
     // Eleminate "third" coordinate
     CASE #pathPlane OF
       "CP_XY":
         #tempVectorA.z := 0.0;
         #tempVectorB.z := 0.0;

       "CP_XZ":
         #tempVectorA.y := 0.0;
         #tempVectorB.y := 0.0;

       "CP_YZ":
         #tempVectorA.x := 0.0;
         #tempVectorB.x := 0.0;
     END_CASE;

     #distancePathPlane := "LKinCtrl_VecAbs"("LKinCtrl_VecSub"(vIn1:=#tempVectorB, vIn2:=#tempVectorA));



   END_REGION CALCULATION

   #LKinCtrl_CalcVecDistancePathPlane := 0; // o.k.
END_FUNCTION

FUNCTION "LKinCtrl_CalcToolLengthCompensation" : Word   // FC35070, SCL
TITLE = LKinCtrl_CalcToolLengthCompensation
{ S7_Optimized_Access := 'TRUE' }
AUTHOR : tech.team.motioncontrol@siemens.com
FAMILY : LKinCtrl
VERSION : 1.0
// Calculate tool length compensation according to path plane and absolute / relative
   VAR_INPUT
      toolLength : LReal;   // Tool length
      pathPlane : Int;   // Path plane: XZ= 0, YZ=1, XY= 2
   END_VAR
   VAR_IN_OUT
      point : "LKinCtrl_typeCOff3DPoint";   // PositioningAxis to get data from
   END_VAR
   // Ret_Val : Return value
   VAR CONSTANT
      ERR_COFF_INVALID_PATH_PLANE : Word := 16#8303;   // Error - invalid path plane
   END_VAR
BEGIN
   //=============================================================================
   // SIEMENS AG
   // (c)Copyright 2019 All Rights Reserved
   //-----------------------------------------------------------------------------
   // Library: - 
   // Tested with: S7-1516T-3 PN
   // Engineering: TIA Portal V15
   // Restrictions: -
   // Requirements: S7-1500/S7-1500T FW 2.5
   // Functionality: Calculate tool length compensation according to path plane and absolute / relative
   // Result ist the compensated coordinate
   // and end point
   //-----------------------------------------------------------------------------
   // Change log table:
   // Version  Date       Expert in charge Changes applied
   // 01.00.00 2019-02-11 AW               created
   //=============================================================================

   REGION PLAUSIBILITY_CHECK
   // Check path plane
   IF ((#pathPlane >= "CP_XZ") AND (#pathPlane <= "CP_XY"))
   THEN
     ;
   ELSE
     #LKinCtrl_CalcToolLengthCompensation := #ERR_COFF_INVALID_PATH_PLANE; // Invalid path plane
     RETURN;
   END_IF;
   END_REGION PLAUSIBILITY_CHECK

   REGION CALCULATION

     CASE #pathPlane OF
       "CP_XY":
         #point.z += #toolLength;
       "CP_XZ":
         #point.y += #toolLength;
       "CP_YZ":
         #point.x += #toolLength;
     END_CASE;


   END_REGION CALCULATION

   #LKinCtrl_CalcToolLengthCompensation := 0; // o.k.
END_FUNCTION

FUNCTION "LKinCtrl_VecAdd" : "LKinCtrl_typeCOff3DPoint"   // FC35080, SCL
TITLE = LKinCtrl_VecAdd
{ S7_Optimized_Access := 'TRUE' }
AUTHOR : tech.team.motioncontrol@siemens.com
FAMILY : LKinCtrl
VERSION : 1.0
// Add two coordinates (X, Y, Z) of "LKinCtrl_typeCOff3DPoint"
   VAR_INPUT
      vIn1 : "LKinCtrl_typeCOff3DPoint";   // Input vector 1
      vIn2 : "LKinCtrl_typeCOff3DPoint";   // Input vector 2
   END_VAR
   // Ret_Val : Return value - calculated vector
BEGIN
   //=============================================================================
   // SIEMENS AG
   // (c)Copyright 2018 All Rights Reserved
   //-----------------------------------------------------------------------------
   // Library: - 
   // Tested with: S7-1516T-3 PN
   // Engineering: TIA Portal V15
   // Restrictions: -
   // Requirements: S7-1500/S7-1500T FW 2.5
   // Functionality: Add two coordinates (X, Y, Z) of "LKinCtrl_typeCOff3DPoint"
   //-----------------------------------------------------------------------------
   // Change log table:
   // Version  Date       Expert in charge Changes applied
   // 01.00.00 2018-10-26 AW               created
   //=============================================================================
   #LKinCtrl_VecAdd.x := #vIn1.x + #vIn2.x;
   #LKinCtrl_VecAdd.y := #vIn1.y + #vIn2.y;
   #LKinCtrl_VecAdd.z := #vIn1.z + #vIn2.z;
END_FUNCTION

FUNCTION "LKinCtrl_VecSub" : "LKinCtrl_typeCOff3DPoint"   // FC35081, SCL
TITLE = LKinCtrl_VecSub
{ S7_Optimized_Access := 'TRUE' }
AUTHOR : tech.team.motioncontrol@siemens.com
FAMILY : LKinCtrl
VERSION : 1.0
// Substract two coordinates (X, Y, Z) of "LKinCtrl_typeCOff3DPoint"
   VAR_INPUT
      vIn1 : "LKinCtrl_typeCOff3DPoint";   // Input vector 1
      vIn2 : "LKinCtrl_typeCOff3DPoint";   // Input vector 2
   END_VAR
   // Ret_Val : Return value - difference vector
BEGIN
   //=============================================================================
   // SIEMENS AG
   // (c)Copyright 2018 All Rights Reserved
   //-----------------------------------------------------------------------------
   // Library: - 
   // Tested with: S7-1516T-3 PN
   // Engineering: TIA Portal V15
   // Restrictions: -
   // Requirements: S7-1500/S7-1500T FW 2.5
   // Functionality: Substract two coordinates (X, Y, Z) of "LKinCtrl_typeCOff3DPoint"
   //-----------------------------------------------------------------------------
   // Change log table:
   // Version  Date       Expert in charge Changes applied
   // 01.00.00 2018-10-26 AW               created
   //=============================================================================
   #LKinCtrl_VecSub.x := #vIn1.x - #vIn2.x;
   #LKinCtrl_VecSub.y := #vIn1.y - #vIn2.y;
   #LKinCtrl_VecSub.z := #vIn1.z - #vIn2.z;
END_FUNCTION

FUNCTION "LKinCtrl_VecUnit" : "LKinCtrl_typeCOff3DPoint"   // FC35082, SCL
TITLE = LKinCtrl_VecUnit
{ S7_Optimized_Access := 'TRUE' }
AUTHOR : tech.team.motioncontrol@siemens.com
FAMILY : LKinCtrl
VERSION : 1.0
// Create unit vector of coordinates (X, Y, Z) of "LKinCtrl_typeCOff3DPoint"
   VAR_INPUT
      vIn : "LKinCtrl_typeCOff3DPoint";   // Input vector
   END_VAR
   // Ret_Val : Return value - unit vector
BEGIN
   //=============================================================================
   // SIEMENS AG
   // (c)Copyright 2018 All Rights Reserved
   //-----------------------------------------------------------------------------
   // Library: - 
   // Tested with: S7-1516T-3 PN
   // Engineering: TIA Portal V15
   // Restrictions: -
   // Requirements: S7-1500/S7-1500T FW 2.5
   // Functionality: Create unit vector of coordinates (X, Y, Z) of "LKinCtrl_typeCOff3DPoint"
   //-----------------------------------------------------------------------------
   // Change log table:
   // Version  Date       Expert in charge Changes applied
   // 01.00.00 2018-08-27 SF               created
   //=============================================================================

   //Out = In/abs(In)
   #LKinCtrl_VecUnit := "LKinCtrl_VecDivScal"(vIn := #vIn,
                                              sIn := "LKinCtrl_VecAbs"(#vIn));
END_FUNCTION

FUNCTION "LKinCtrl_VecAbs" : LReal   // FC35083, SCL
TITLE = LKinCtrl_VecAbs
{ S7_Optimized_Access := 'TRUE' }
AUTHOR : tech.team.motioncontrol@siemens.com
FAMILY : LKinCtrl
VERSION : 1.0
// Calculate length of vector of coordinates (X, Y, Z) of "LKinCtrl_typeCOff3DPoint"
   VAR_INPUT
      vIn : "LKinCtrl_typeCOff3DPoint";   // Input vector
   END_VAR
   // Ret_Val : Return value - scalar
BEGIN
   //=============================================================================
   // SIEMENS AG
   // (c)Copyright 2018 All Rights Reserved
   //-----------------------------------------------------------------------------
   // Library: - 
   // Tested with: S7-1516T-3 PN
   // Engineering: TIA Portal V15
   // Restrictions: -
   // Requirements: S7-1500/S7-1500T FW 2.5
   // Functionality: Calculate length of vector of coordinates (X, Y, Z) of "LKinCtrl_typeCOff3DPoint"
   //-----------------------------------------------------------------------------
   // Change log table:
   // Version  Date       Expert in charge Changes applied
   // 01.00.00 2018-10-26 AW               created
   //=============================================================================

   #LKinCtrl_VecAbs := SQRT(#vIn.x*#vIn.x + #vIn.y*#vIn.y + #vIn.z*#vIn.z);
END_FUNCTION

FUNCTION "LKinCtrl_VecScale" : "LKinCtrl_typeCOff3DPoint"   // FC35084, SCL
TITLE = LKinCtrl_VecScale
{ S7_Optimized_Access := 'TRUE' }
AUTHOR : tech.team.motioncontrol@siemens.com
FAMILY : LKinCtrl
VERSION : 1.0
// Scale vector (X, Y, Z) of "LKinCtrl_typeCOff3DPoint"
   VAR_INPUT
      vIn : "LKinCtrl_typeCOff3DPoint";   // Input vector
      factor : LReal;   // Scaling factor
   END_VAR
   // Ret_Val : Return value - scaled vector
BEGIN
   //=============================================================================
   // SIEMENS AG
   // (c)Copyright 2018 All Rights Reserved
   //-----------------------------------------------------------------------------
   // Library: - 
   // Tested with: S7-1516T-3 PN
   // Engineering: TIA Portal V15
   // Restrictions: -
   // Requirements: S7-1500/S7-1500T FW 2.5
   // Functionality: Scale vector (X, Y, Z) of "LKinCtrl_typeCOff3DPoint"
   //-----------------------------------------------------------------------------
   // Change log table:
   // Version  Date       Expert in charge Changes applied
   // 01.00.00 2018-10-26 AW               created
   //=============================================================================

   #LKinCtrl_VecScale.x := #vIn.x * #factor;
   #LKinCtrl_VecScale.y := #vIn.y * #factor;
   #LKinCtrl_VecScale.z := #vIn.z * #factor;
END_FUNCTION

FUNCTION "LKinCtrl_VecDivScal" : "LKinCtrl_typeCOff3DPoint"   // FC35085, SCL
TITLE = LKinCtrl_VecDivScal
{ S7_Optimized_Access := 'TRUE' }
AUTHOR : tech.team.motioncontrol@siemens.com
FAMILY : LKinCtrl
VERSION : 1.0
// Divide coordinate with scalar of coordinates (X, Y, Z) of "LKinCtrl_typeCOff3DPoint"
   VAR_INPUT
      vIn : "LKinCtrl_typeCOff3DPoint";   // Input vector
      sIn : LReal;   // Input scalar
   END_VAR
   // Ret_Val : Return value - calculated vector
BEGIN
   //=============================================================================
   // SIEMENS AG
   // (c)Copyright 2018 All Rights Reserved
   //-----------------------------------------------------------------------------
   // Library: - 
   // Tested with: S7-1516T-3 PN
   // Engineering: TIA Portal V15
   // Restrictions: -
   // Requirements: S7-1500/S7-1500T FW 2.5
   // Functionality: Divide coordinate with scalar of coordinates (X, Y, Z) of "LKinCtrl_typeCOff3DPoint"
   //-----------------------------------------------------------------------------
   // Change log table:
   // Version  Date       Expert in charge Changes applied
   // 01.00.00 2018-10-26 AW               created
   //=============================================================================

   IF (#sIn <> 0.0) THEN
     #LKinCtrl_VecDivScal.x := #vIn.x / #sIn;
     #LKinCtrl_VecDivScal.y := #vIn.y / #sIn;
     #LKinCtrl_VecDivScal.z := #vIn.z / #sIn;
   ELSE
     #LKinCtrl_VecDivScal.x := 0.0;
     #LKinCtrl_VecDivScal.y := 0.0;
     #LKinCtrl_VecDivScal.z := 0.0;
   END_IF;
END_FUNCTION

FUNCTION "LKinCtrl_VecScalProd" : LReal   // FC35086, SCL
TITLE = LKinCtrl_VecScalProd
{ S7_Optimized_Access := 'TRUE' }
AUTHOR : tech.team.motioncontrol@siemens.com
FAMILY : LKinCtrl
VERSION : 1.0
// Calculate scalar product of coordinates (X, Y, Z) of "LKinCtrl_typeCOff3DPoint"
   VAR_INPUT
      vIn1 : "LKinCtrl_typeCOff3DPoint";   // Input vector 1
      vIn2 : "LKinCtrl_typeCOff3DPoint";   // Input vector 2
   END_VAR
   // Ret_Val : Scalar product
BEGIN
   //=============================================================================
   // SIEMENS AG
   // (c)Copyright 2019 All Rights Reserved
   //-----------------------------------------------------------------------------
   // Library: - 
   // Tested with: S7-1516T-3 PN
   // Engineering: TIA Portal V15
   // Restrictions: -
   // Requirements: S7-1500/S7-1500T FW 2.5
   // Functionality: Calculate scalar product of coordinates (X, Y, Z) of "LKinCtrl_typeCOff3DPoint"
   //-----------------------------------------------------------------------------
   // Change log table:
   // Version  Date       Expert in charge Changes applied
   // 01.00.00 2019-01-25 AW               created
   //=============================================================================

   #LKinCtrl_VecScalProd := #vIn1.x * #vIn2.x  //   X1*X2
                          + #vIn1.y * #vIn2.y  // + Y1*Y2
                          + #vIn1.z * #vIn2.z; // + Z1*Z2
END_FUNCTION

FUNCTION "LKinCtrl_VecCrossProd" : "LKinCtrl_typeCOff3DPoint"   // FC35087, SCL
TITLE = LKinCtrl_VecCrossProd
{ S7_Optimized_Access := 'TRUE' }
AUTHOR : tech.team.motioncontrol@siemens.com
FAMILY : LKinCtrl
VERSION : 1.0
// Cross product of two coordinates (X, Y, Z) of "LKinCtrl_typeCOff3DPoint"
   VAR_INPUT
      vIn1 : "LKinCtrl_typeCOff3DPoint";   // Input vector 1
      vIn2 : "LKinCtrl_typeCOff3DPoint";   // Input vector 2
   END_VAR
   // Ret_Val : Return value - calculated vector
BEGIN
   //=============================================================================
   // SIEMENS AG
   // (c)Copyright 2018 All Rights Reserved
   //-----------------------------------------------------------------------------
   // Library: - 
   // Tested with: S7-1516T-3 PN
   // Engineering: TIA Portal V15
   // Restrictions: -
   // Requirements: S7-1500/S7-1500T FW 2.5
   // Functionality: Cross product of two coordinates (X, Y, Z) of "LKinCtrl_typeCOff3DPoint"
   //-----------------------------------------------------------------------------
   // Change log table:
   // Version  Date       Expert in charge Changes applied
   // 01.00.00 2019-01-24 AW               created
   //=============================================================================

   #LKinCtrl_VecCrossProd.x := #vIn1.y * #vIn2.z - #vIn1.z * #vIn2.y;
   #LKinCtrl_VecCrossProd.y := #vIn1.z * #vIn2.x - #vIn1.x * #vIn2.z;
   #LKinCtrl_VecCrossProd.z := #vIn1.x * #vIn2.y - #vIn1.y * #vIn2.x;
END_FUNCTION

// folder: LKinCtrl_Blocks/LKinCtrl_SubBlocks/LKinCtrl_SubCalcBlocks

FUNCTION_BLOCK "LKinCtrl_SetFlagCtrl"   // FB35024, SCL
TITLE = LKinCtrl_SetFlagCtrl / Enable Template
{ S7_Optimized_Access := 'TRUE' }
AUTHOR : tech.team.motioncontrol@siemens.com
FAMILY : LKinCtrl
VERSION : 2.0
// Handle setFlags in FB MovePath / Template for an FB with Enable / Valid handling based on PLCopen standard "Function Blocks for Motion Control" V2.0
   VAR_INPUT
      enable : Bool;   // TRUE: Enable functionality of FB
      activeCmdNo : DInt;   // Number of actual PathData set number (interconnect LKinCtrl_MC_ExecuteKinMotionCmd)
      activePathDataIdentifier : USInt;   // Identifier number of actual PathData (interconnect LKinCtrl_MC_ExecuteKinMotionCmd)
      activePathDataName : String["LKINCTRL_LENGTH_OF_PATHDATA_NAME"];   // Name of actual PathData (interconnect LKinCtrl_MC_ExecuteKinMotionCmd)
      remainingDistanceActCmd : LReal;   // RemainingDistance of active motionCommand (interconnect LKinCtrl_MC_ExecuteKinMotionCmd)
      kinematicsStatusWord : DWord;   // Interconnect axesGroup.StatusWord / Interconnect 'axesGroup.StatusWord.X9'
      movePathStatus : Word;   // Interconnect value for MovePath output 'status'
      flagsBuffer : Struct   // Buffer to store flag information for past and actual commands
         writeBufferElement : Int := 1;   // pointer on entry to be written
         bufferElement : Array[1.."LKINCTRL_NO_OF_SETFLAGS_BUFFER_ELEMENTS"] of Struct   // flag information for one specific command (see cmdId)
            pathDataName : String["LKINCTRL_LENGTH_OF_PATHDATA_NAME"];   // PathData name of specific command
            pathDataIdentifier : DInt;   // PathData identifier counter of specific command
            cmdId : DInt;   // cmdId of command in PathData
            isIntermediateCmd : Bool;   // TRUE: command is intermediate command
            setFlags : Array[1.."LKINCTRL_NO_OF_CMD_SETFLAGS"] of "LKinCtrl_typeSetFlagElement_Bool";   // setFlags structure equal to PathData command entry
            valueFlags : Array[1.."LKINCTRL_NO_OF_CMD_VALUEFLAGS"] of "LKinCtrl_typeSetFlagElement_LReal";   // setFlags structure equal to PathData command entry
         END_STRUCT;
      END_STRUCT;
   END_VAR
   VAR_OUTPUT
      valid : Bool;   // TRUE: Valid set of output values available at the FB
      busy : Bool;   // TRUE: FB is not finished and new output values can be expected
      error : Bool;   // TRUE: An error occurred during the execution of the FB
      status : Word := 16#7000;   // 16#0000 - 16#7FFF: Status of the FB, 16#8000 - 16#FFFF: Error identification
      waitMain : Bool;   // Static bit to wait for execution due to wait flags & valueFlags
   END_VAR
   VAR_IN_OUT
      flags : Array[0.."LKINCTRL_NO_OF_LAST_SETFLAG"] of Bool;   // Interconnect MovePath outputs for flag signals
      waitFlags : Struct   // Static struct to store wait flag information
         waitCtr : Int;   // counter for number of wait flags in one command
         waitFlag : Array[1.."LKINCTRL_NO_OF_CMD_SETFLAGS"] of Int;   // flag number as identifier for flag active as wait flag
      END_STRUCT;
   END_VAR
   VAR
      statEnableOld : Bool;   // Old value of 'enable' input for edge detection
      statValid : Bool;   // Static value for output 'valid'
      statBusy : Bool;   // Static value for output 'busy'
      statError : Bool;   // Static value for output 'error'
      statErrorUserCleared : Bool;   // Error occurred that can only be solved by user; rising edge at enable input necessary
      statErrorAutoCleared : Bool;   // Error occurred that can be acknowledged by FB
      statStatus : Word := 16#7000;   // Static value for output 'status'
      statFBState : DInt := 0;   // State in the state machine of the FB
      statDisablingCompleted : Bool;   // TRUE: Disabling has been completed
      statWaitMain : Bool;   // Static value for output 'waitMain'
      statSkippedCmdCounter : Int;   // Static counter for skipped activeCmdNo
      statActivePathDataIdentifierOld : USInt;   // Static to store old activePathDataIdentifier from LKinCtrl_ExecuteKinMotionCmd
      statActiveCmdNoOld : DInt;   // Static variable storing old 'activeCmdNo'
      statActivePathDataNameOld : String["LKINCTRL_LENGTH_OF_PATHDATA_NAME"];   // Static to store last active PathData name
      statFlagSetAfterCmd : Array[1.."LKINCTRL_NO_OF_CMD_SETFLAGS"] of Int;   // Static array storing flags to be set after command
      statWaitFlagSetAfterCmd : Array[1.."LKINCTRL_NO_OF_CMD_SETFLAGS"] of Int;   // Static array storing wait flags to be set after command / Static array storing flags to be set after command
      statFlagResetAfterOneCmd : Array[1.."LKINCTRL_NO_OF_CMD_SETFLAGS"] of Int;   // Static array storing flags to be reset after one command
      statFlagResetFM3 : Array[1.."LKINCTRL_NO_OF_CMD_SETFLAGS"] of Int;   // Static array storing flags to be reset after one cycle
      statFlagSetFM10 : Array[1.."LKINCTRL_NO_OF_CMD_SETFLAGS"] of Int;   // Static array storing flags to be set at remaining distance
      statRemDistanceFM10 : Array[1.."LKINCTRL_NO_OF_CMD_SETFLAGS"] of LReal;   // Static array storing remaining distance for flags
      statFlagSetFM13 : Array[1.."LKINCTRL_NO_OF_CMD_SETFLAGS"] of Int;   // Static array storing flags to be set after command for one cycle
      statFlagResetFM13 : Array[1.."LKINCTRL_NO_OF_CMD_SETFLAGS"] of Int;   // Static array storing flags to be set after command and reset after one cycle
      statWaitFlagActiveCmdId : Array[1.."LKINCTRL_NO_OF_CMD_SETFLAGS"] of DInt;   // Static array storing active command number for watiFlag
      statWaitFlagActivePathData : Array[1.."LKINCTRL_NO_OF_CMD_SETFLAGS"] of DInt;   // Static array storing active PathData number for watiFlag
      statFlagResetSkipped : Array[1..#MAX_NUMBER_OF_SKIPPED_CMDS, 1.."LKINCTRL_NO_OF_CMD_SETFLAGS"] of Int;   // Static array storing flags to be reset after one cycle
      statWaitFlagOld : Array[1.."LKINCTRL_NO_OF_CMD_SETFLAGS"] of Bool;   // Static array storing last flag values for reset detection
   END_VAR
   VAR_TEMP
      tempEnable : Bool;   // Temporary value for input 'enable'
      tempFlagCmdCounter : Int;   // Temporary flag cmd counter for setFlag UDT
      tempFlagsBufferElementCtr : Int;   // Temporary flag buffer counter
      tempFlagCounter : Int;   // Temporary flag counter for flag array
      tempFlagWasSet : Bool;   // Temporary bool to signalize flag was set after end of PRG
      tempSkippedCounterInc : Bool;   // Temporary bool to signalize skipped counter was increased
   END_VAR
   VAR CONSTANT
      FB_STATE_NO_PROCESSING : DInt := 0;   // FB state: No processing
      FB_STATE_CHECK_ACTIVE_CMD : DInt := 50;   // FB state: Check change of active command
      FB_STATE_SET_RESET_AFTER_COMMAND : DInt := 51;   // FB state: Handle flag actions after commands
      FB_STATE_EVALUATE_FLAGBUFFER : DInt := 52;   // FB state: Handle flagBuffer and flag actions before command
      FB_STATE_RESET_AFTER_ONE_CYCLE : DInt := 53;   // FB state: Handle flag reset after one cycle
      FB_STATE_CHECK_REMAINING_DISTANCE : DInt := 54;   // FB state: Check flag with remaining distance
      FB_STATE_WAIT_FLAG_HANDLING : DInt := 55;   // FB state: Check wait flags
      FB_STATE_DISABLING : DInt := 90;   // FB state: Disabling
      STATUS_NO_CALL : Word := 16#7000;   // No job being currently processed
      STATUS_FIRST_CALL : Word := 16#7001;   // First call after incoming new job (rising edge 'execute')
      STATUS_SUBSEQUENT_CALL : Word := 16#7002;   // Subsequent call during active processing without further details
      ERR_UNDEFINED_STATE : Word := 16#8600;   // Error due to an undefined state in state machine
      ERR_OVERFLOW_SKIPPED_CMDS : Word := 16#8601;   // Error due to overflow of skipped commands counter
      STATUS_EXECUTION_WAITING : Word := 16#7307;   // Status path execution waiting due to wait flag, wait time or single step mode
      MAX_NUMBER_OF_SKIPPED_CMDS : Int := 3;   // Maximum number of activeCmdNo to be skipped
      SPTP_REMAINING_DIST : Bool := FALSE;   // TRUE: Caclulate own RemainingDistance for SPTP / FALSE: Use ExecutionTimeStatus
   END_VAR
   // flagsBuffer.bufferElement[1].pathDataName := '';
   // flagsBuffer.bufferElement[1].cmdId := 0;
BEGIN
   //==========================================================================================
   // SIEMENS AG
   // (c)Copyright 2020 All Rights Reserved
   //------------------------------------------------------------------------------------------
   // Library: LKinCtrl
   // Tested with: S7-1517T-3 PN/DP
   // Engineering: TIA Portal V15
   // Restrictions: ---
   // Requirements: S7-1500T FW 2.5
   // Functionality: LKinCtrl_SetFlagCtrl
   // The FC evaluates the flag informaton given by the PathData structure and controls the flag
   // variables depending on the active command information given
   // 
   // Support: tech.team.motioncontrol@siemens.com
   // Note: Parameter comments are only available in language 'English (United States)'
   //------------------------------------------------------------------------------------------
   // Change log table:
   // Version    Date          Expert in charge    Changes applied
   // 01.00.00   19.08.2019    JR                  First release version v1.0
   // 01.00.01   18.09.2019    JR                  Updates for LREAL flags
   // 01.00.02   19.09.2019    JR                  Implementation wait value flags - flagMode 5
   // 01.00.03   19.09.2019    JR                  Implementation value flags - flagMode 11 - 15
   // 01.00.04   27.11.2019    JR                  Additional condition for deactivating flags
   // 01.01.00   28.11.2019    JR                  Separate block for setFlags from LKinCtrl_FlagCtrl
   // 01.01.01   27.01.2020    FR                  Changed FM 10 from > to >=
   // 01.01.02   30.01.2020    FR                  Changed flag array constant
   // 02.00.00   12.03.2020    FR                  Reworked complete FB to fit enable template with state machine
   // 02.00.01   17.03.2020    FR                  Check remDistance <= 0.0 instead of =
   // 02.00.02   03.08.2020    FR                  Change interface actualCmdIsCircularCmd to KinematicsStatusWord (DWord)
   // 02.00.03   19.10.2020    FR                  Handle multiple commands per cycle; Changed case to use constants instead of numbers
   // 02.00.04   15.12.2020    FR                  Added option for SPTP commands to have calculated remainingDistance
   // 02.00.05   01.06.2021    FR                  Use variable instead of F_Trig, Fix for FM5 / FM15, Fix for statActiveCmdNoOld not being reset correctly
   // 02.00.06   06.07.2021    FR                  Save old variables only when processed
   //===========================================================================================

   #tempEnable := #enable; // Work with temporary value / create process image

   REGION ENABLING/DISABLING
     IF (#tempEnable = TRUE) AND (#statStatus = #STATUS_NO_CALL) THEN // Enable FB
       // First call; initialize FB
       #statValid := TRUE;
       #statBusy := TRUE;
       #statError := FALSE;
       #statErrorUserCleared := FALSE;
       #statErrorAutoCleared := FALSE;
       #statStatus := #STATUS_FIRST_CALL;

       #statFBState := #FB_STATE_CHECK_ACTIVE_CMD; // State machine - start functionality
       //------------------------------------------------------------------------------------------
       // Initialize functionality: reset of variables, diagnostics, etc.
       #statDisablingCompleted := FALSE;

       // Initialize all setFlags (flag array) when enabling
       //------------------------------------------------------------------------------------------
       FOR #tempFlagCounter := 0 TO "LKINCTRL_NO_OF_LAST_SETFLAG" DO
         #flags[#tempFlagCounter] := FALSE;
       END_FOR;

       // Initialize flag handling variables
       //------------------------------------------------------------------------------------------
       // reset wait output
       #statWaitMain := FALSE;
       #statSkippedCmdCounter := 0;
       #statActiveCmdNoOld := 0;
       #statActivePathDataNameOld := '';
       #statActivePathDataIdentifierOld := 0;

       FOR #tempFlagCmdCounter := 1 TO "LKINCTRL_NO_OF_CMD_SETFLAGS" DO
         // reset auxiliary flag storage variables
         #statFlagResetAfterOneCmd[#tempFlagCmdCounter] := -1;
         #statFlagSetAfterCmd[#tempFlagCmdCounter] := -1;
         #statWaitFlagSetAfterCmd[#tempFlagCmdCounter] := -1;
         #statFlagResetFM3[#tempFlagCmdCounter] := -1;
         #statFlagResetFM13[#tempFlagCmdCounter] := -1;
         #statFlagSetFM13[#tempFlagCmdCounter] := -1;
         #statFlagSetFM10[#tempFlagCmdCounter] := -1;
         #statRemDistanceFM10[#tempFlagCmdCounter] := 0.0;
         #statWaitFlagActiveCmdId[#tempFlagCmdCounter] := 0;
         #statWaitFlagActivePathData[#tempFlagCmdCounter] := 0;

         // Initialize functionality: call subsidiary FBs with FALSE
         #statWaitFlagOld[#tempFlagCmdCounter] := FALSE;

         // Reset storage for skipped commands
         FOR #tempFlagCounter := 1 TO #MAX_NUMBER_OF_SKIPPED_CMDS DO
           #statFlagResetSkipped[#tempFlagCounter, #tempFlagCmdCounter] := -1;
         END_FOR;
       END_FOR;


       //------------------------------------------------------------------------------------------

     ELSIF (#tempEnable = FALSE) AND (#statEnableOld = TRUE) THEN // Disable FB 
       #statFBState := #FB_STATE_DISABLING;

     ELSIF (#statStatus = #STATUS_FIRST_CALL) THEN // Set status identifier of subsequent call
       #statStatus := #STATUS_SUBSEQUENT_CALL;
     END_IF;

     // Edge detection 'enable' input
     #statEnableOld := #tempEnable;
   END_REGION ENABLING/DISABLING

   IF (#statStatus = #STATUS_NO_CALL) THEN // Nothing to do -> End here to reduce "system load"
     RETURN;
   END_IF;

   REGION STATE_MACHINE
     // Use if sate machine for more states in one cycle

     // No processing active (Note: this state must always be present and left empty)
     IF #statFBState = #FB_STATE_NO_PROCESSING THEN
       ;
     END_IF;

     // Reset after one cycle 
     REGION STATE_RESET_AFTER_ONE_CYCLE
       IF #statFBState = #FB_STATE_RESET_AFTER_ONE_CYCLE THEN
         // for loop checking all available flags
         FOR #tempFlagCmdCounter := 1 TO "LKINCTRL_NO_OF_CMD_SETFLAGS" DO
           // reset flags active for one cycle only (flagMode: 3)
           IF #statFlagResetFM3[#tempFlagCmdCounter] <> -1 THEN
             // reset flags when active command is ended / next command starts
             #flags[#statFlagResetFM3[#tempFlagCmdCounter]] := FALSE;
             // reset stored flag to be reset (to not reset it after each single future command)
             #statFlagResetFM3[#tempFlagCmdCounter] := -1;
           END_IF;

           // reset flags active for one cycle only (flagMode: 13)
           IF #statFlagResetFM13[#tempFlagCmdCounter] <> -1 THEN
             // reset flags when active command is ended / next command starts
             #flags[#statFlagResetFM13[#tempFlagCmdCounter]] := FALSE;
             // reset stored flag to be reset (to not reset it after each single future command)
             #statFlagResetFM13[#tempFlagCmdCounter] := -1;
           END_IF;

           // Check if commands were skipped and reset flags
           FOR #tempFlagCounter := 1 TO #statSkippedCmdCounter DO // If no cmd was skipped the upper limit should be 0 --> No execution of the loop
             // If activeCmdNo was skipped reset flags active for one cycle only (flagMode: 2/3/13)
             IF #statFlagResetSkipped[#tempFlagCounter, #tempFlagCmdCounter] <> -1 THEN
               // reset flags when active command is ended / next command starts
               #flags[#statFlagResetSkipped[#tempFlagCounter, #tempFlagCmdCounter]] := FALSE;
               // reset stored flag to be reset (to not reset it after each single future command)
               #statFlagResetSkipped[#tempFlagCounter, #tempFlagCmdCounter] := -1;
             END_IF;
           END_FOR;
         END_FOR;

         // go to next state
         #statFBState := #FB_STATE_CHECK_ACTIVE_CMD;
       END_IF;
     END_REGION STATE_RESET_AFTER_ONE_CYCLE


     // Cyclic state
     // This state shall be the idle state where conditions are checked 
     // --> Change in active command number
     // --> End of cmd
     // --> End of prg
     // --> ...
     REGION STATE_CHECK_ACTIVE_CMD
       IF #statFBState = #FB_STATE_CHECK_ACTIVE_CMD THEN // Processing active
         // Check if activeCmdNo has changed or MovePath is waiting and remainingDistance = 0
         // --> Go to state: #FB_STATE_SET_RESET_AFTER_COMMAND
         // Else
         // --> Go to state: #FB_STATE_CHECK_REMAINING_DISTANCE
         // 
         // Check if active cmd no has changed // changed JR 2019/04/11 < to <>
         IF (#statActiveCmdNoOld <> #activeCmdNo OR #statActivePathDataIdentifierOld <> #activePathDataIdentifier)
           OR (#movePathStatus = #STATUS_EXECUTION_WAITING AND #remainingDistanceActCmd <= 0.0) // check for command to be finished
         THEN
           #statFBState := #FB_STATE_SET_RESET_AFTER_COMMAND;
         ELSE
           #statFBState := #FB_STATE_CHECK_REMAINING_DISTANCE;
         END_IF;
       END_IF;
     END_REGION STATE_CHECK_ACTIVE_CMD


     // Set / Reset flags after command has finished (FM2 / FM11 / FM13 / FM15)
     REGION STATE_SET_RESET_AFTER_COMMAND
       IF #statFBState = #FB_STATE_SET_RESET_AFTER_COMMAND THEN
         // for loop checking all available flags
         FOR #tempFlagCmdCounter := 1 TO "LKINCTRL_NO_OF_CMD_SETFLAGS" DO
           // reset flags active for one command only (flagMode: 2 (LKINCTRL_FM_SET_BEFORE_AND_RESET_AFTER))
           IF #statFlagResetAfterOneCmd[#tempFlagCmdCounter] <> -1 THEN
             // reset flags when active command is ended / next command starts
             #flags[#statFlagResetAfterOneCmd[#tempFlagCmdCounter]] := FALSE;
             // reset stored flag to be reset (to not reset it after each single future command)
             #statFlagResetAfterOneCmd[#tempFlagCmdCounter] := -1;
           END_IF;

           // set flags to be activated at end of command
           // flagMode: 11 (LKINCTRL_FM_SET_AFTER_AND_NO_RESET)
           IF #statFlagSetAfterCmd[#tempFlagCmdCounter] <> -1 THEN
             // set flags when active command is ended / next command starts
             #flags[#statFlagSetAfterCmd[#tempFlagCmdCounter]] := TRUE;
             // reset stored flag to be set (to not set it after each single future command)
             #statFlagSetAfterCmd[#tempFlagCmdCounter] := -1;
           END_IF;

           // flagMode: 15 (LKINCTRL_FM_SET_AFTER_AND_NO_RESET_AND_WAIT_FOR_ACKNOWLEDGE)
           IF #statWaitFlagSetAfterCmd[#tempFlagCmdCounter] <> -1 THEN
             // set flags when active command is ended / next command starts
             #flags[#statWaitFlagSetAfterCmd[#tempFlagCmdCounter]] := TRUE;
             #statWaitFlagOld[#tempFlagCmdCounter] := TRUE;
             // reset stored flag to be set (to not set it after each single future command)
             #statWaitFlagSetAfterCmd[#tempFlagCmdCounter] := -1;
           END_IF;

           // set flags to be activated at end of command
           // flagMode: 13 (LKINCTRL_FM_SET_AFTER_AND_RESET_AFTER_ONE_CYCLE)
           IF #statFlagSetFM13[#tempFlagCmdCounter] <> -1 THEN
             // set flags when active command is ended / next command starts
             #flags[#statFlagSetFM13[#tempFlagCmdCounter]] := TRUE;

             // Save flag numbers to be reset after one cycle
             #statFlagResetFM13[#tempFlagCmdCounter] := #statFlagSetFM13[#tempFlagCmdCounter];

             // reset stored flag to be set (to not set it after each single future command)
             #statFlagSetFM13[#tempFlagCmdCounter] := -1;
           END_IF;

           // Check if FM10 was not executed and set if next command is reached
           IF (#statFlagSetFM10[#tempFlagCmdCounter] <> -1) THEN
             // Set flag if remaining distance is reached
             #flags[#statFlagSetFM10[#tempFlagCmdCounter]] := TRUE;
             // reset stored flag to be reset (to not reset it after each single future command)
             #statFlagSetFM10[#tempFlagCmdCounter] := -1;
             #statRemDistanceFM10[#tempFlagCmdCounter] := 0.0;
           END_IF;

         END_FOR;

         // go to next state ; skip new flag if waiting
         IF #movePathStatus = #STATUS_EXECUTION_WAITING
           AND NOT (#statActiveCmdNoOld <> #activeCmdNo OR #statActivePathDataIdentifierOld <> #activePathDataIdentifier)
         THEN
           #statFBState := #FB_STATE_CHECK_REMAINING_DISTANCE;
         ELSE
           #statFBState := #FB_STATE_EVALUATE_FLAGBUFFER;
         END_IF;
       END_IF;
     END_REGION STATE_SET_RESET_AFTER_COMMAND

     // Set flags before command and save variables to set after command (STATE_SET_RESET_AFTER)
     // This state shall be used to copy flag buffer into variables 
     // This state is reached after the state to set/reset flags after a command 
     // --> Set flags before command instantly 
     // --> Set flags after command in next call because of the state machine order
     REGION STATE_EVALUATE_FLAGBUFFER
       IF #statFBState = #FB_STATE_EVALUATE_FLAGBUFFER THEN
         // Reset counter
         #statSkippedCmdCounter := 0;

         // Reset activeCmdNoOld when PathData changes
         IF #activeCmdNo = 1 THEN
           #statActiveCmdNoOld := 0;
         END_IF;

         // only run flag controls when a set is active
         IF #activeCmdNo > 0 THEN
           // selection of active flags and evaluation of flagMode
           FOR #tempFlagsBufferElementCtr := 1 TO "LKINCTRL_NO_OF_SETFLAGS_BUFFER_ELEMENTS" DO
             IF #flagsBuffer.bufferElement[#tempFlagsBufferElementCtr].pathDataIdentifier = #activePathDataIdentifier // choose correct setFlags stored according to corresponding PathData
               AND #flagsBuffer.bufferElement[#tempFlagsBufferElementCtr].cmdId <= #activeCmdNo // choose only flags to be controlled when corresponding command is active
               AND #flagsBuffer.bufferElement[#tempFlagsBufferElementCtr].cmdId > #statActiveCmdNoOld // Also check flags on previous commands
             THEN
               // Reset temp to allow skippedCmdCounter to be increased
               #tempSkippedCounterInc := FALSE;

               // set flags according to PathData configuration stored in #statStoreSetFlagsBuffer
               FOR #tempFlagCmdCounter := 1 TO "LKINCTRL_NO_OF_CMD_SETFLAGS" DO

                 // check for flag not to be deactivated
                 IF #flagsBuffer.bufferElement[#tempFlagsBufferElementCtr].setFlags[#tempFlagCmdCounter].flag > -1 THEN

                   CASE #flagsBuffer.bufferElement[#tempFlagsBufferElementCtr].setFlags[#tempFlagCmdCounter].flagMode OF
                       //------------------------------------------------------------------------------------------
                     "LKINCTRL_FM_SET_BEFORE_AND_NO_RESET": // FM 1
                       // (activate flag at beginning of command)
                       // set selected flag to TRUE at beginning of command
                       #flags[#flagsBuffer.bufferElement[#tempFlagsBufferElementCtr].setFlags[#tempFlagCmdCounter].flag] := TRUE;
                       //------------------------------------------------------------------------------------------

                       //------------------------------------------------------------------------------------------
                     "LKINCTRL_FM_SET_BEFORE_AND_RESET_AFTER": // FM 2
                       // (activate flag at beginning of command)
                       // set selected flag to TRUE at beginning of command
                       #flags[#flagsBuffer.bufferElement[#tempFlagsBufferElementCtr].setFlags[#tempFlagCmdCounter].flag] := TRUE;

                       IF #flagsBuffer.bufferElement[#tempFlagsBufferElementCtr].cmdId = #activeCmdNo THEN
                         // store flags to be set for one command only to reset at the end of command
                         #statFlagResetAfterOneCmd[#tempFlagCmdCounter] := #flagsBuffer.bufferElement[#tempFlagsBufferElementCtr].setFlags[#tempFlagCmdCounter].flag;
                       ELSE
                         // Check if skippedCmdCounter must be increased
                         IF NOT #tempSkippedCounterInc THEN
                           #statSkippedCmdCounter += 1;
                           #tempSkippedCounterInc := TRUE; // Store bit to avoid counting several times per command
                           IF #statSkippedCmdCounter > #MAX_NUMBER_OF_SKIPPED_CMDS THEN
                             // Throw error
                             #statStatus := #ERR_OVERFLOW_SKIPPED_CMDS;
                             #statErrorUserCleared := TRUE;
                             EXIT;
                           END_IF;
                         END_IF;
                         // ActiveCmdNo was skipped --> Store flag number to be reset after one cycle
                         #statFlagResetSkipped[#statSkippedCmdCounter, #tempFlagCmdCounter] := #flagsBuffer.bufferElement[#tempFlagsBufferElementCtr].setFlags[#tempFlagCmdCounter].flag;
                       END_IF;
                       //------------------------------------------------------------------------------------------

                       //------------------------------------------------------------------------------------------
                     "LKINCTRL_FM_SET_BEFORE_AND_RESET_AFTER_ONE_CYCLE": // FM 3
                       // (activate flag at beginning of command for one cycle only)
                       // set selected flag to TRUE at beginning of command
                       #flags[#flagsBuffer.bufferElement[#tempFlagsBufferElementCtr].setFlags[#tempFlagCmdCounter].flag] := TRUE;

                       IF #flagsBuffer.bufferElement[#tempFlagsBufferElementCtr].cmdId = #activeCmdNo THEN
                         #statFlagResetFM3[#tempFlagCmdCounter] := #flagsBuffer.bufferElement[#tempFlagsBufferElementCtr].setFlags[#tempFlagCmdCounter].flag;
                       ELSE
                         // Check if skippedCmdCounter must be increased
                         IF NOT #tempSkippedCounterInc THEN
                           #statSkippedCmdCounter += 1;
                           #tempSkippedCounterInc := TRUE; // Store bit to avoid counting several times per command
                           IF #statSkippedCmdCounter > #MAX_NUMBER_OF_SKIPPED_CMDS THEN
                             // Throw error
                             #statStatus := #ERR_OVERFLOW_SKIPPED_CMDS;
                             #statErrorUserCleared := TRUE;
                             EXIT;
                           END_IF;
                         END_IF;
                         // ActiveCmdNo was skipped --> Store flag number to be reset after one cycle
                         #statFlagResetSkipped[#statSkippedCmdCounter, #tempFlagCmdCounter] := #flagsBuffer.bufferElement[#tempFlagsBufferElementCtr].setFlags[#tempFlagCmdCounter].flag;
                       END_IF;
                       //------------------------------------------------------------------------------------------

                       //------------------------------------------------------------------------------------------ 
                     "LKINCTRL_FM_SET_BEFORE_AND_NO_RESET_AND_WAIT_FOR_ACKNOWLEDGE": // FM 5
                       // (activate flag at beginning of command and continue path motion only after acknowledge (reset) of set flag)
                       #flags[#flagsBuffer.bufferElement[#tempFlagsBufferElementCtr].setFlags[#tempFlagCmdCounter].flag] := TRUE;
                       #statWaitFlagOld[#tempFlagCmdCounter] := TRUE;
                       // Store active command information for edge detection
                       // --> Avoid edge detection in wrong command
                       #statWaitFlagActiveCmdId[#tempFlagCmdCounter] := #activeCmdNo;
                       #statWaitFlagActivePathData[#tempFlagCmdCounter] := #activePathDataIdentifier;
                       //------------------------------------------------------------------------------------------ 

                     "LKINCTRL_FM_SET_AT_REMAINING_DISTANCE": // FM 10
                       // FM 10 is checked cyclic
                       IF #flagsBuffer.bufferElement[#tempFlagsBufferElementCtr].cmdId = #activeCmdNo THEN
                         #statFlagSetFM10[#tempFlagCmdCounter] := #flagsBuffer.bufferElement[#tempFlagsBufferElementCtr].setFlags[#tempFlagCmdCounter].flag;
                         #statRemDistanceFM10[#tempFlagCmdCounter] := #flagsBuffer.bufferElement[#tempFlagsBufferElementCtr].setFlags[#tempFlagCmdCounter].remainingDistance;
                       ELSE
                         // ActiveCmdNo was skipped --> Set flag instantly
                         #flags[#flagsBuffer.bufferElement[#tempFlagsBufferElementCtr].setFlags[#tempFlagCmdCounter].flag] := TRUE;
                       END_IF;

                       //------------------------------------------------------------------------------------------
                     "LKINCTRL_FM_SET_AFTER_AND_NO_RESET": // FM 11
                       // activate flag at end of command
                       IF #flagsBuffer.bufferElement[#tempFlagsBufferElementCtr].cmdId = #activeCmdNo THEN
                         // store flags to be set at the end of command and not being reset
                         #statFlagSetAfterCmd[#tempFlagCmdCounter] := #flagsBuffer.bufferElement[#tempFlagsBufferElementCtr].setFlags[#tempFlagCmdCounter].flag;
                       ELSE
                         // ActiveCmdNo was skipped --> Set flag instantly
                         #flags[#flagsBuffer.bufferElement[#tempFlagsBufferElementCtr].setFlags[#tempFlagCmdCounter].flag] := TRUE;
                       END_IF;
                       //------------------------------------------------------------------------------------------

                       //------------------------------------------------------------------------------------------
                     "LKINCTRL_FM_SET_AFTER_AND_RESET_AFTER_ONE_CYCLE": // FM 13
                       // activate flag at end of command
                       IF #flagsBuffer.bufferElement[#tempFlagsBufferElementCtr].cmdId = #activeCmdNo THEN
                         // store flags to be set at the end of command and to be reset after one cycle
                         #statFlagSetFM13[#tempFlagCmdCounter] := #flagsBuffer.bufferElement[#tempFlagsBufferElementCtr].setFlags[#tempFlagCmdCounter].flag;
                       ELSE
                         // ActiveCmdNo was skipped --> Set flag instantly and reset after one cycle
                         #flags[#flagsBuffer.bufferElement[#tempFlagsBufferElementCtr].setFlags[#tempFlagCmdCounter].flag] := TRUE;
                         // Check if skippedCmdCounter must be increased
                         IF NOT #tempSkippedCounterInc THEN
                           #statSkippedCmdCounter += 1;
                           #tempSkippedCounterInc := TRUE; // Store bit to avoid counting several times per command
                           IF #statSkippedCmdCounter > #MAX_NUMBER_OF_SKIPPED_CMDS THEN
                             // Throw error
                             #statStatus := #ERR_OVERFLOW_SKIPPED_CMDS;
                             #statErrorUserCleared := TRUE;
                             EXIT;
                           END_IF;
                         END_IF;
                         // ActiveCmdNo was skipped --> Store flag number to be reset after one cycle
                         #statFlagResetSkipped[#statSkippedCmdCounter, #tempFlagCmdCounter] := #flagsBuffer.bufferElement[#tempFlagsBufferElementCtr].setFlags[#tempFlagCmdCounter].flag;
                       END_IF;
                       //------------------------------------------------------------------------------------------

                       //------------------------------------------------------------------------------------------
                     "LKINCTRL_FM_SET_AFTER_AND_NO_RESET_AND_WAIT_FOR_ACKNOWLEDGE": // FM 15
                       // activate flag at end of command and continue path motion only after acknowledge (reset) of set flag
                       // store flags to be set at the end of command and not being reset
                       #statWaitFlagSetAfterCmd[#tempFlagCmdCounter] := #flagsBuffer.bufferElement[#tempFlagsBufferElementCtr].setFlags[#tempFlagCmdCounter].flag;
                       // Store active command information for edge detection
                       // --> Avoid edge detection in wrong command
                       #statWaitFlagActiveCmdId[#tempFlagCmdCounter] := #activeCmdNo;
                       #statWaitFlagActivePathData[#tempFlagCmdCounter] := #activePathDataIdentifier;
                       //------------------------------------------------------------------------------------------

                     ELSE
                       ;
                   END_CASE;
                 END_IF;
               END_FOR;
             END_IF;

             // In case of error also exit outer loop
             IF #statErrorUserCleared THEN
               EXIT;
             END_IF;

           END_FOR;

           // Save "old" variables
           #statActiveCmdNoOld := #activeCmdNo;
           #statActivePathDataNameOld := #activePathDataName;
           #statActivePathDataIdentifierOld := #activePathDataIdentifier;
         END_IF;

         // go to next state 
         #statFBState := #FB_STATE_CHECK_REMAINING_DISTANCE;
       END_IF;
     END_REGION STATE_EVALUATE_FLAGBUFFER

     // Check remaining distance of actual command for FM10 (LKINCTRL_FM_SET_AT_REMAINING_DISTANCE)
     REGION STATE_CHECK_REMAINING_DISTANCE
       IF #statFBState = #FB_STATE_CHECK_REMAINING_DISTANCE THEN
         FOR #tempFlagCmdCounter := 1 TO "LKINCTRL_NO_OF_CMD_SETFLAGS" DO
           // Set flags in remaining distance FM10
           IF (#statFlagSetFM10[#tempFlagCmdCounter] <> -1)
             AND (((#remainingDistanceActCmd <= #statRemDistanceFM10[#tempFlagCmdCounter])
             AND (#kinematicsStatusWord.%X11 = FALSE)) // No SPTP active
             OR ((#remainingDistanceActCmd >= #statRemDistanceFM10[#tempFlagCmdCounter])
             AND (#kinematicsStatusWord.%X11 = TRUE) AND (#SPTP_REMAINING_DIST = FALSE)) // SPTP active, regular
             OR ((#remainingDistanceActCmd <= #statRemDistanceFM10[#tempFlagCmdCounter])
             AND (#kinematicsStatusWord.%X11 = TRUE) AND (#SPTP_REMAINING_DIST = TRUE))) // SPTP active, remDistance calculated
           THEN
             // Set flag if remaining distance is reached
             #flags[#statFlagSetFM10[#tempFlagCmdCounter]] := TRUE;
             // reset stored flag to be reset (to not reset it after each single future command)
             #statFlagSetFM10[#tempFlagCmdCounter] := -1;
             #statRemDistanceFM10[#tempFlagCmdCounter] := 0.0;
           END_IF;
         END_FOR;

         // Go to next state
         #statFBState := #FB_STATE_WAIT_FLAG_HANDLING;
       END_IF;
     END_REGION STATE_CHECK_REMAINING_DISTANCE

